// TIA Portal project "SMSS-ENLAB-01-003-1508-012-PLC-B_V13_SP1_1_V17" (V17) (continued)
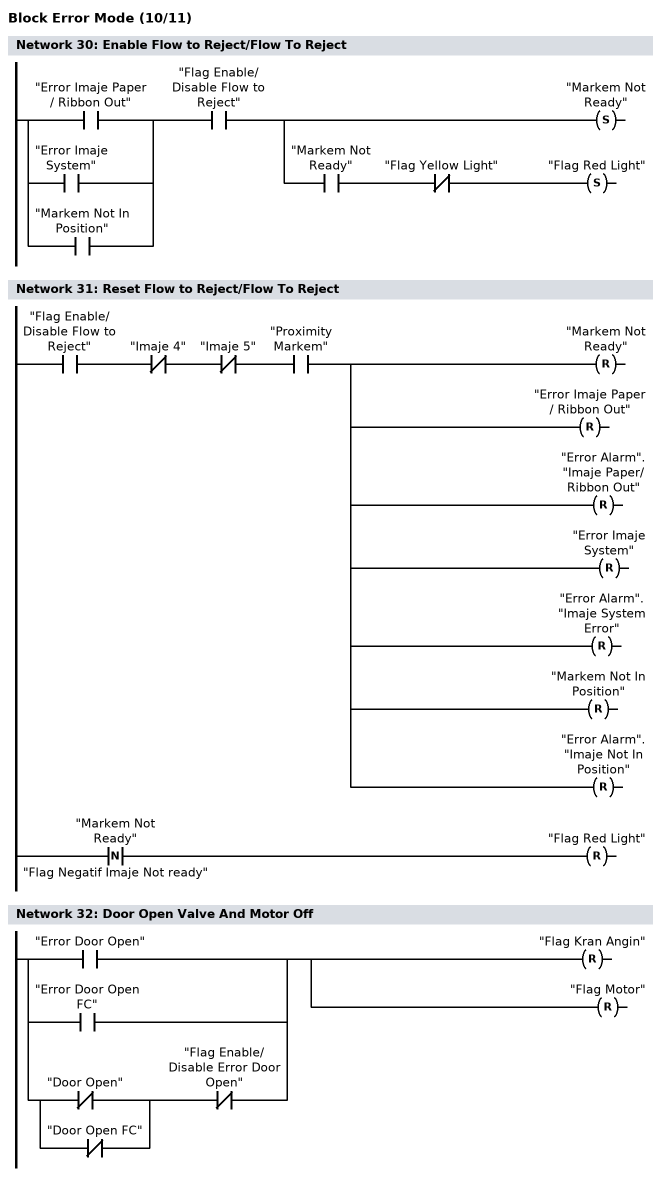
   RUNG wire#powerrail
      Contact( "Error Imaje Paper / Ribbon Out" )
      wire#w1
      Contact( "Flag Enable/Disable Flow to Reject" )
      wire#w2
      S_Coil( "Markem Not Ready" )
   END_RUNG
   RUNG wire#powerrail
      Contact( "Error Imaje System" )
   END_RUNG wire#w1
   RUNG wire#powerrail
      Contact( "Markem Not In Position" )
   END_RUNG wire#w1
   RUNG wire#w2
      Contact( "Markem Not Ready" )
      I_Contact( "Flag Yellow Light" )
      S_Coil( "Flag Red Light" )
   END_RUNG
   // the same network as SCL:
   #_w1 := ("Error Imaje Paper / Ribbon Out" OR "Error Imaje System" OR "Markem Not In Position") AND "Flag Enable/Disable Flow to Reject";
   IF #_w1 THEN "Markem Not Ready" := TRUE; END_IF;
   IF #_w1 AND "Markem Not Ready" AND NOT "Flag Yellow Light" THEN "Flag Red Light" := TRUE; END_IF;
END_REGION

REGION Network 31: Reset Flow to Reject/Flow To Reject
   RUNG wire#powerrail
      Contact( "Flag Enable/Disable Flow to Reject" )
      I_Contact( "Imaje 4" )
      I_Contact( "Imaje 5" )
      Contact( "Proximity Markem" )
      wire#w1
      R_Coil( "Markem Not Ready" )
   END_RUNG
   RUNG wire#w1
      R_Coil( "Error Imaje Paper / Ribbon Out" )
   END_RUNG
   RUNG wire#w1
      R_Coil( "Error Alarm"."Imaje Paper/Ribbon Out" )
   END_RUNG
   RUNG wire#w1
      R_Coil( "Error Imaje System" )
   END_RUNG
   RUNG wire#w1
      R_Coil( "Error Alarm"."Imaje System Error" )
   END_RUNG
   RUNG wire#w1
      R_Coil( "Markem Not In Position" )
   END_RUNG
   RUNG wire#w1
      R_Coil( "Error Alarm"."Imaje Not In Position" )
   END_RUNG
   RUNG wire#powerrail
      N_Contact(operand := "Markem Not Ready", bit := "Flag Negatif Imaje Not ready")
      R_Coil( "Flag Red Light" )
   END_RUNG
   // the same network as SCL:
   IF "Flag Enable/Disable Flow to Reject" AND NOT "Imaje 4" AND NOT "Imaje 5" AND "Proximity Markem" THEN
       "Markem Not Ready" := FALSE;
       "Error Imaje Paper / Ribbon Out" := FALSE;
       "Error Alarm"."Imaje Paper/Ribbon Out" := FALSE;
       "Error Imaje System" := FALSE;
       "Error Alarm"."Imaje System Error" := FALSE;
       "Markem Not In Position" := FALSE;
       "Error Alarm"."Imaje Not In Position" := FALSE;
   END_IF;
   #_w1 := NOT "Markem Not Ready" AND "Flag Negatif Imaje Not ready";   // falling edge of "Markem Not Ready"
   "Flag Negatif Imaje Not ready" := "Markem Not Ready";
   IF #_w1 THEN "Flag Red Light" := FALSE; END_IF;
END_REGION

REGION Network 32: Door Open Valve And Motor Off
   RUNG wire#powerrail
      Contact( "Error Door Open" )
      wire#w1
      R_Coil( "Flag Kran Angin" )
   END_RUNG
   RUNG wire#powerrail
      Contact( "Error Door Open FC" )
   END_RUNG wire#w1
   RUNG wire#powerrail
      I_Contact( "Door Open" )
      wire#w2
      I_Contact( "Flag Enable/Disable Error Door Open" )
   END_RUNG wire#w1
   RUNG wire#powerrail
      I_Contact( "Door Open FC" )
   END_RUNG wire#w2
   RUNG wire#w1
      R_Coil( "Flag Motor" )
   END_RUNG
   // the same network as SCL:
   IF "Error Door Open" OR "Error Door Open FC" OR ((NOT "Door Open" OR NOT "Door Open FC") AND NOT "Flag Enable/Disable Error Door Open") THEN
       "Flag Kran Angin" := FALSE;
       "Flag Motor" := FALSE;
   END_IF;
END_REGION

REGION Network 33: Baypas Error Reset error 3
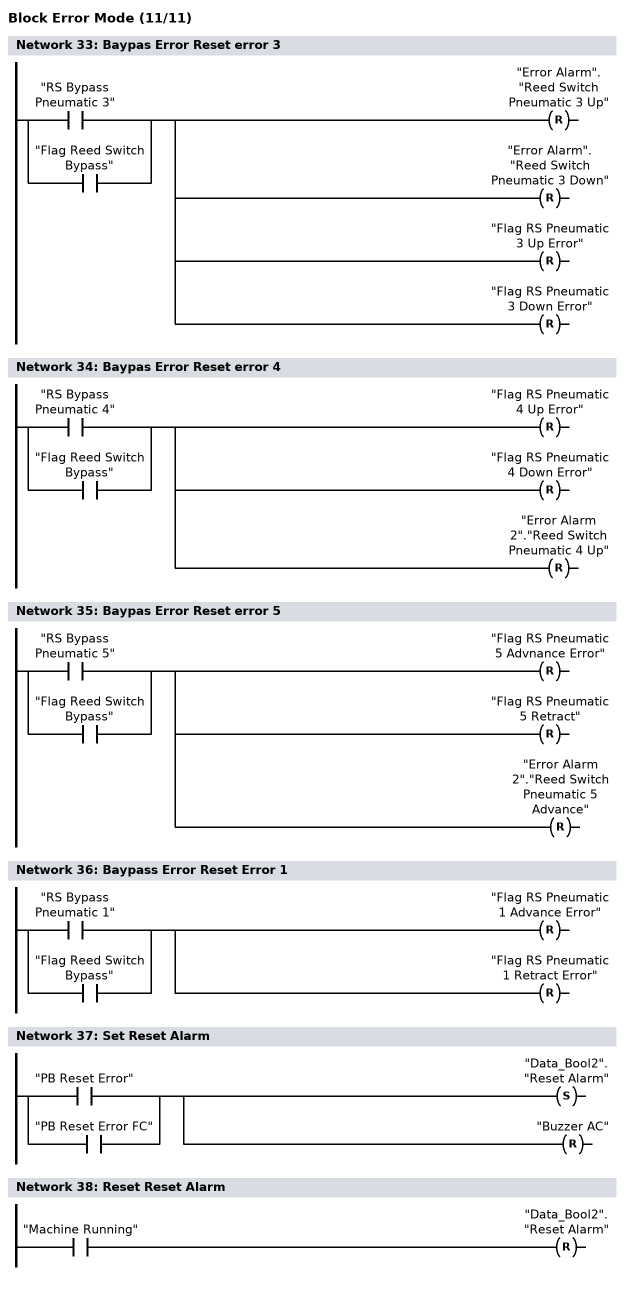
   RUNG wire#powerrail
      Contact( "RS Bypass Pneumatic 3" )
      wire#w1
      R_Coil( "Error Alarm"."Reed Switch Pneumatic 3 Up" )
   END_RUNG
   RUNG wire#powerrail
      Contact( "Flag Reed Switch Bypass" )
   END_RUNG wire#w1
   RUNG wire#w1
      R_Coil( "Error Alarm"."Reed Switch Pneumatic 3 Down" )
   END_RUNG
   RUNG wire#w1
      R_Coil( "Flag RS Pneumatic 3 Up Error" )
   END_RUNG
   RUNG wire#w1
      R_Coil( "Flag RS Pneumatic 3 Down Error" )
   END_RUNG
   // the same network as SCL:
   IF "RS Bypass Pneumatic 3" OR "Flag Reed Switch Bypass" THEN
       "Error Alarm"."Reed Switch Pneumatic 3 Up" := FALSE;
       "Error Alarm"."Reed Switch Pneumatic 3 Down" := FALSE;
       "Flag RS Pneumatic 3 Up Error" := FALSE;
       "Flag RS Pneumatic 3 Down Error" := FALSE;
   END_IF;
END_REGION

REGION Network 34: Baypas Error Reset error 4
   RUNG wire#powerrail
      Contact( "RS Bypass Pneumatic 4" )
      wire#w1
      R_Coil( "Flag RS Pneumatic 4 Up Error" )
   END_RUNG
   RUNG wire#powerrail
      Contact( "Flag Reed Switch Bypass" )
   END_RUNG wire#w1
   RUNG wire#w1
      R_Coil( "Flag RS Pneumatic 4 Down Error" )
   END_RUNG
   RUNG wire#w1
      R_Coil( "Error Alarm 2"."Reed Switch Pneumatic 4 Up" )
   END_RUNG
   // the same network as SCL:
   IF "RS Bypass Pneumatic 4" OR "Flag Reed Switch Bypass" THEN
       "Flag RS Pneumatic 4 Up Error" := FALSE;
       "Flag RS Pneumatic 4 Down Error" := FALSE;
       "Error Alarm 2"."Reed Switch Pneumatic 4 Up" := FALSE;
   END_IF;
END_REGION

REGION Network 35: Baypas Error Reset error 5
   RUNG wire#powerrail
      Contact( "RS Bypass Pneumatic 5" )
      wire#w1
      R_Coil( "Flag RS Pneumatic 5 Advnance Error" )
   END_RUNG
   RUNG wire#powerrail
      Contact( "Flag Reed Switch Bypass" )
   END_RUNG wire#w1
   RUNG wire#w1
      R_Coil( "Flag RS Pneumatic 5 Retract" )
   END_RUNG
   RUNG wire#w1
      R_Coil( "Error Alarm 2"."Reed Switch Pneumatic 5 Advance" )
   END_RUNG
   // the same network as SCL:
   IF "RS Bypass Pneumatic 5" OR "Flag Reed Switch Bypass" THEN
       "Flag RS Pneumatic 5 Advnance Error" := FALSE;
       "Flag RS Pneumatic 5 Retract" := FALSE;
       "Error Alarm 2"."Reed Switch Pneumatic 5 Advance" := FALSE;
   END_IF;
END_REGION

REGION Network 36: Baypass Error Reset Error 1
   RUNG wire#powerrail
      Contact( "RS Bypass Pneumatic 1" )
      wire#w1
      R_Coil( "Flag RS Pneumatic 1 Advance Error" )
   END_RUNG
   RUNG wire#powerrail
      Contact( "Flag Reed Switch Bypass" )
   END_RUNG wire#w1
   RUNG wire#w1
      R_Coil( "Flag RS Pneumatic 1 Retract Error" )
   END_RUNG
   // the same network as SCL:
   IF "RS Bypass Pneumatic 1" OR "Flag Reed Switch Bypass" THEN
       "Flag RS Pneumatic 1 Advance Error" := FALSE;
       "Flag RS Pneumatic 1 Retract Error" := FALSE;
   END_IF;
END_REGION

REGION Network 37: Set Reset Alarm
   RUNG wire#powerrail
      Contact( "PB Reset Error" )
      wire#w1
      S_Coil( "Data_Bool2"."Reset Alarm" )
   END_RUNG
   RUNG wire#powerrail
      Contact( "PB Reset Error FC" )
   END_RUNG wire#w1
   RUNG wire#w1
      R_Coil( "Buzzer AC" )
   END_RUNG
   // the same network as SCL:
   IF "PB Reset Error" OR "PB Reset Error FC" THEN
       "Data_Bool2"."Reset Alarm" := TRUE;
       "Buzzer AC" := FALSE;
   END_IF;
END_REGION

REGION Network 38: Reset Reset Alarm
   RUNG wire#powerrail
      Contact( "Machine Running" )
      R_Coil( "Data_Bool2"."Reset Alarm" )
   END_RUNG
   // the same network as SCL:
   IF "Machine Running" THEN "Data_Bool2"."Reset Alarm" := FALSE; END_IF;
END_REGION
END_FUNCTION_BLOCK

FUNCTION_BLOCK "Block Test Mode"   // FB2, LAD
{ S7_Optimized_Access := 'TRUE' }
VERSION : 0.1
BEGIN

REGION Network 1: Set Motor Conveyor
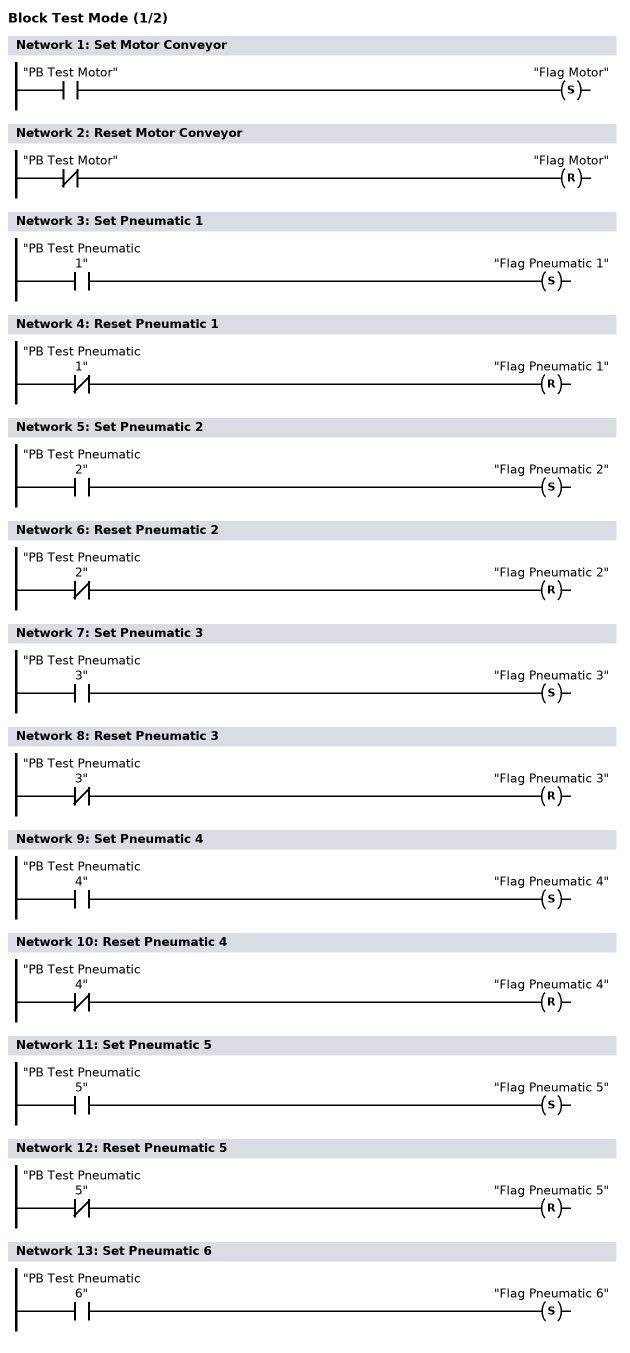
   RUNG wire#powerrail
      Contact( "PB Test Motor" )
      S_Coil( "Flag Motor" )
   END_RUNG
   // the same network as SCL:
   IF "PB Test Motor" THEN "Flag Motor" := TRUE; END_IF;
END_REGION

REGION Network 2: Reset Motor Conveyor
   RUNG wire#powerrail
      I_Contact( "PB Test Motor" )
      R_Coil( "Flag Motor" )
   END_RUNG
   // the same network as SCL:
   IF NOT "PB Test Motor" THEN "Flag Motor" := FALSE; END_IF;
END_REGION

REGION Network 3: Set Pneumatic 1
   RUNG wire#powerrail
      Contact( "PB Test Pneumatic 1" )
      S_Coil( "Flag Pneumatic 1" )
   END_RUNG
   // the same network as SCL:
   IF "PB Test Pneumatic 1" THEN "Flag Pneumatic 1" := TRUE; END_IF;
END_REGION

REGION Network 4: Reset Pneumatic 1
   RUNG wire#powerrail
      I_Contact( "PB Test Pneumatic 1" )
      R_Coil( "Flag Pneumatic 1" )
   END_RUNG
   // the same network as SCL:
   IF NOT "PB Test Pneumatic 1" THEN "Flag Pneumatic 1" := FALSE; END_IF;
END_REGION

REGION Network 5: Set Pneumatic 2
   RUNG wire#powerrail
      Contact( "PB Test Pneumatic 2" )
      S_Coil( "Flag Pneumatic 2" )
   END_RUNG
   // the same network as SCL:
   IF "PB Test Pneumatic 2" THEN "Flag Pneumatic 2" := TRUE; END_IF;
END_REGION

REGION Network 6: Reset Pneumatic 2
   RUNG wire#powerrail
      I_Contact( "PB Test Pneumatic 2" )
      R_Coil( "Flag Pneumatic 2" )
   END_RUNG
   // the same network as SCL:
   IF NOT "PB Test Pneumatic 2" THEN "Flag Pneumatic 2" := FALSE; END_IF;
END_REGION

REGION Network 7: Set Pneumatic 3
   RUNG wire#powerrail
      Contact( "PB Test Pneumatic 3" )
      S_Coil( "Flag Pneumatic 3" )
   END_RUNG
   // the same network as SCL:
   IF "PB Test Pneumatic 3" THEN "Flag Pneumatic 3" := TRUE; END_IF;
END_REGION

REGION Network 8: Reset Pneumatic 3
   RUNG wire#powerrail
      I_Contact( "PB Test Pneumatic 3" )
      R_Coil( "Flag Pneumatic 3" )
   END_RUNG
   // the same network as SCL:
   IF NOT "PB Test Pneumatic 3" THEN "Flag Pneumatic 3" := FALSE; END_IF;
END_REGION

REGION Network 9: Set Pneumatic 4
   RUNG wire#powerrail
      Contact( "PB Test Pneumatic 4" )
      S_Coil( "Flag Pneumatic 4" )
   END_RUNG
   // the same network as SCL:
   IF "PB Test Pneumatic 4" THEN "Flag Pneumatic 4" := TRUE; END_IF;
END_REGION

REGION Network 10: Reset Pneumatic 4
   RUNG wire#powerrail
      I_Contact( "PB Test Pneumatic 4" )
      R_Coil( "Flag Pneumatic 4" )
   END_RUNG
   // the same network as SCL:
   IF NOT "PB Test Pneumatic 4" THEN "Flag Pneumatic 4" := FALSE; END_IF;
END_REGION

REGION Network 11: Set Pneumatic 5
   RUNG wire#powerrail
      Contact( "PB Test Pneumatic 5" )
      S_Coil( "Flag Pneumatic 5" )
   END_RUNG
   // the same network as SCL:
   IF "PB Test Pneumatic 5" THEN "Flag Pneumatic 5" := TRUE; END_IF;
END_REGION

REGION Network 12: Reset Pneumatic 5
   RUNG wire#powerrail
      I_Contact( "PB Test Pneumatic 5" )
      R_Coil( "Flag Pneumatic 5" )
   END_RUNG
   // the same network as SCL:
   IF NOT "PB Test Pneumatic 5" THEN "Flag Pneumatic 5" := FALSE; END_IF;
END_REGION

REGION Network 13: Set Pneumatic 6
   RUNG wire#powerrail
      Contact( "PB Test Pneumatic 6" )
      S_Coil( "Flag Pneumatic 6" )
   END_RUNG
   // the same network as SCL:
   IF "PB Test Pneumatic 6" THEN "Flag Pneumatic 6" := TRUE; END_IF;
END_REGION

REGION Network 14: Reset Pneumatic 6
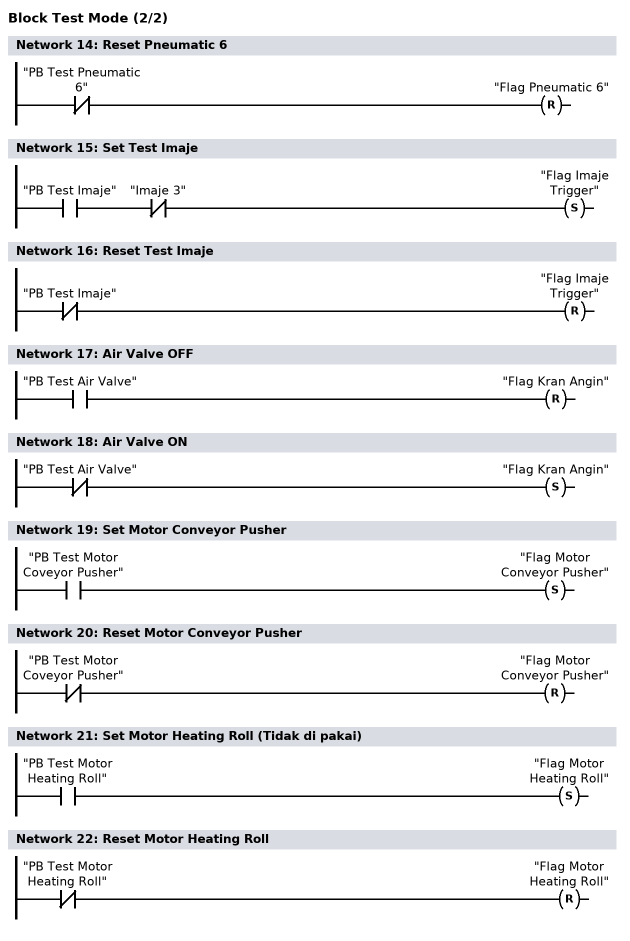
   RUNG wire#powerrail
      I_Contact( "PB Test Pneumatic 6" )
      R_Coil( "Flag Pneumatic 6" )
   END_RUNG
   // the same network as SCL:
   IF NOT "PB Test Pneumatic 6" THEN "Flag Pneumatic 6" := FALSE; END_IF;
END_REGION

REGION Network 15: Set Test Imaje
   RUNG wire#powerrail
      Contact( "PB Test Imaje" )
      I_Contact( "Imaje 3" )
      S_Coil( "Flag Imaje Trigger" )
   END_RUNG
   // the same network as SCL:
   IF "PB Test Imaje" AND NOT "Imaje 3" THEN "Flag Imaje Trigger" := TRUE; END_IF;
END_REGION

REGION Network 16: Reset Test Imaje
   RUNG wire#powerrail
      I_Contact( "PB Test Imaje" )
      R_Coil( "Flag Imaje Trigger" )
   END_RUNG
   // the same network as SCL:
   IF NOT "PB Test Imaje" THEN "Flag Imaje Trigger" := FALSE; END_IF;
END_REGION

REGION Network 17: Air Valve OFF
   RUNG wire#powerrail
      Contact( "PB Test Air Valve" )
      R_Coil( "Flag Kran Angin" )
   END_RUNG
   // the same network as SCL:
   IF "PB Test Air Valve" THEN "Flag Kran Angin" := FALSE; END_IF;
END_REGION

REGION Network 18: Air Valve ON
   RUNG wire#powerrail
      I_Contact( "PB Test Air Valve" )
      S_Coil( "Flag Kran Angin" )
   END_RUNG
   // the same network as SCL:
   IF NOT "PB Test Air Valve" THEN "Flag Kran Angin" := TRUE; END_IF;
END_REGION

REGION Network 19: Set Motor Conveyor Pusher
   RUNG wire#powerrail
      Contact( "PB Test Motor Coveyor Pusher" )
      S_Coil( "Flag Motor Conveyor Pusher" )
   END_RUNG
   // the same network as SCL:
   IF "PB Test Motor Coveyor Pusher" THEN "Flag Motor Conveyor Pusher" := TRUE; END_IF;
END_REGION

REGION Network 20: Reset Motor Conveyor Pusher
   RUNG wire#powerrail
      I_Contact( "PB Test Motor Coveyor Pusher" )
      R_Coil( "Flag Motor Conveyor Pusher" )
   END_RUNG
   // the same network as SCL:
   IF NOT "PB Test Motor Coveyor Pusher" THEN "Flag Motor Conveyor Pusher" := FALSE; END_IF;
END_REGION

REGION Network 21: Set Motor Heating Roll (Tidak di pakai)
   RUNG wire#powerrail
      Contact( "PB Test Motor Heating Roll" )
      S_Coil( "Flag Motor Heating Roll" )
   END_RUNG
   // the same network as SCL:
   IF "PB Test Motor Heating Roll" THEN "Flag Motor Heating Roll" := TRUE; END_IF;
END_REGION

REGION Network 22: Reset Motor Heating Roll
   RUNG wire#powerrail
      I_Contact( "PB Test Motor Heating Roll" )
      R_Coil( "Flag Motor Heating Roll" )
   END_RUNG
   // the same network as SCL:
   IF NOT "PB Test Motor Heating Roll" THEN "Flag Motor Heating Roll" := FALSE; END_IF;
END_REGION
END_FUNCTION_BLOCK

FUNCTION_BLOCK "Block Output"   // FB3, LAD
{ S7_Optimized_Access := 'TRUE' }
VERSION : 0.1
   VAR_TEMP   // added for the SCL form of the ladder/FBD networks
      _w1 : Bool;
      _w2 : Bool;
      _w3 : Bool;
   END_VAR
BEGIN

REGION Network 1: Red Light Tower
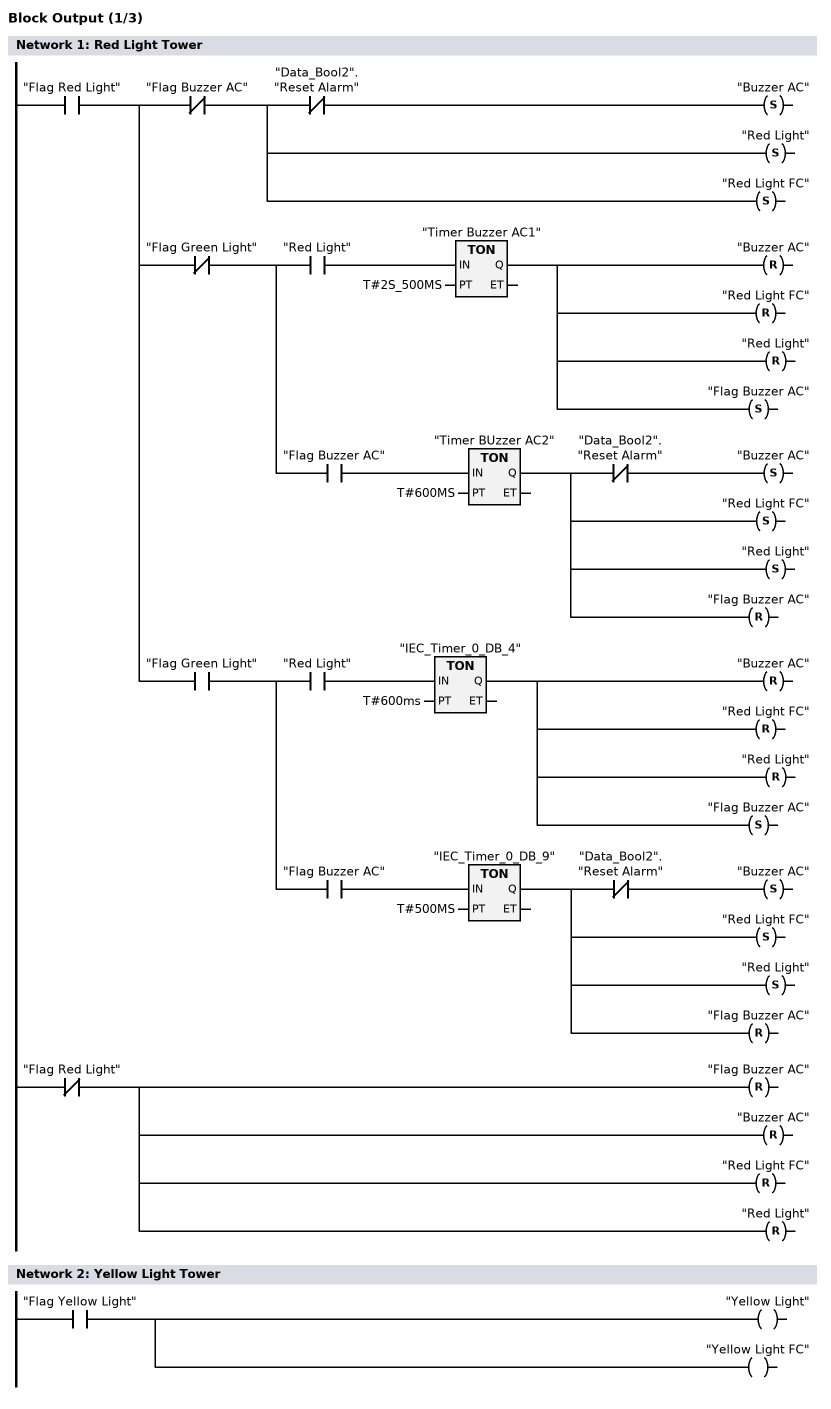
   #_w1 := "Flag Red Light" AND NOT "Flag Buzzer AC";
   IF #_w1 AND NOT "Data_Bool2"."Reset Alarm" THEN "Buzzer AC" := TRUE; END_IF;
   IF #_w1 THEN
       "Red Light" := TRUE;
       "Red Light FC" := TRUE;
   END_IF;
   #_w2 := "Flag Red Light" AND NOT "Flag Green Light";
   "Timer Buzzer AC1".TON(IN := #_w2 AND "Red Light", PT := T#2S_500MS);
   IF "Timer Buzzer AC1".Q THEN
       "Buzzer AC" := FALSE;
       "Red Light FC" := FALSE;
       "Red Light" := FALSE;
       "Flag Buzzer AC" := TRUE;
   END_IF;
   "Timer BUzzer AC2".TON(IN := #_w2 AND "Flag Buzzer AC", PT := T#600MS);
   IF "Timer BUzzer AC2".Q AND NOT "Data_Bool2"."Reset Alarm" THEN "Buzzer AC" := TRUE; END_IF;
   IF "Timer BUzzer AC2".Q THEN
       "Red Light FC" := TRUE;
       "Red Light" := TRUE;
       "Flag Buzzer AC" := FALSE;
   END_IF;
   #_w3 := "Flag Red Light" AND "Flag Green Light";
   "IEC_Timer_0_DB_4".TON(IN := #_w3 AND "Red Light", PT := T#600ms);
   IF "IEC_Timer_0_DB_4".Q THEN
       "Buzzer AC" := FALSE;
       "Red Light FC" := FALSE;
       "Red Light" := FALSE;
       "Flag Buzzer AC" := TRUE;
   END_IF;
   "IEC_Timer_0_DB_9".TON(IN := #_w3 AND "Flag Buzzer AC", PT := T#500MS);
   IF "IEC_Timer_0_DB_9".Q AND NOT "Data_Bool2"."Reset Alarm" THEN "Buzzer AC" := TRUE; END_IF;
   IF "IEC_Timer_0_DB_9".Q THEN
       "Red Light FC" := TRUE;
       "Red Light" := TRUE;
       "Flag Buzzer AC" := FALSE;
   END_IF;
   IF NOT "Flag Red Light" THEN
       "Flag Buzzer AC" := FALSE;
       "Buzzer AC" := FALSE;
       "Red Light FC" := FALSE;
       "Red Light" := FALSE;
   END_IF;
END_REGION

REGION Network 2: Yellow Light Tower
   RUNG wire#powerrail
      Contact( "Flag Yellow Light" )
      wire#w1
      Coil( "Yellow Light" )
   END_RUNG
   RUNG wire#w1
      Coil( "Yellow Light FC" )
   END_RUNG
   // the same network as SCL:
   "Yellow Light" := "Flag Yellow Light";
   "Yellow Light FC" := "Flag Yellow Light";
END_REGION

REGION Network 3: Green Light Tower
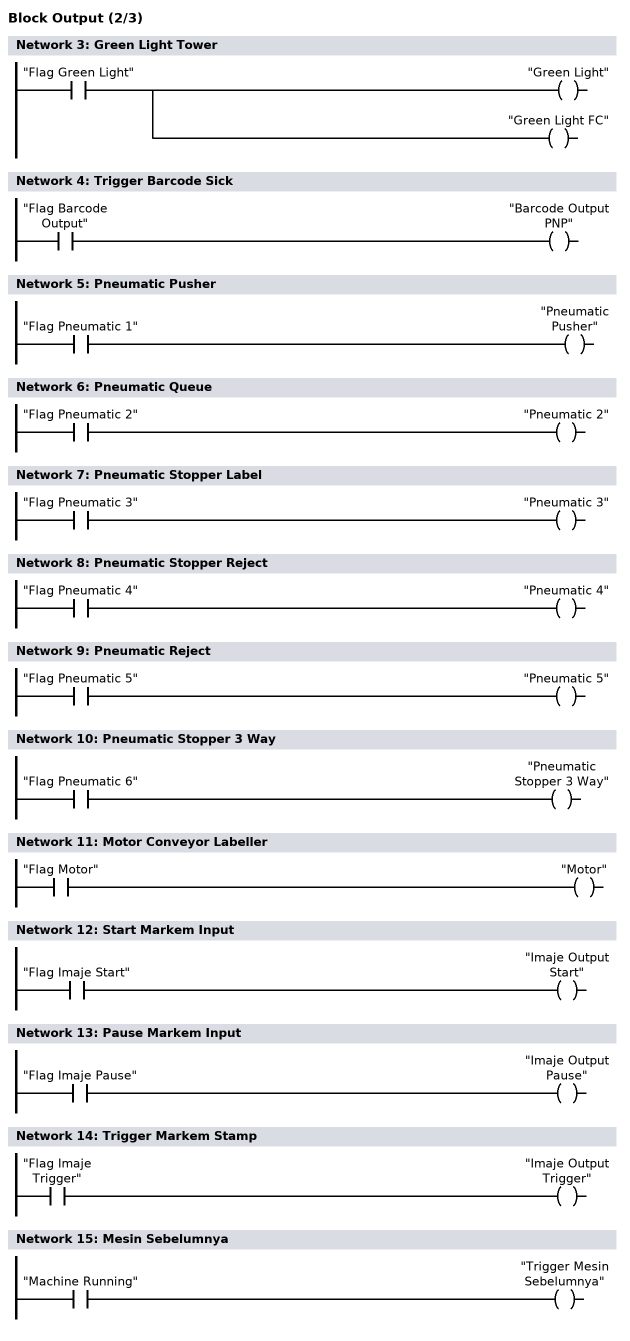
   RUNG wire#powerrail
      Contact( "Flag Green Light" )
      wire#w1
      Coil( "Green Light" )
   END_RUNG
   RUNG wire#w1
      Coil( "Green Light FC" )
   END_RUNG
   // the same network as SCL:
   "Green Light" := "Flag Green Light";
   "Green Light FC" := "Flag Green Light";
END_REGION

REGION Network 4: Trigger Barcode Sick
   RUNG wire#powerrail
      Contact( "Flag Barcode Output" )
      Coil( "Barcode Output PNP" )
   END_RUNG
   // the same network as SCL:
   "Barcode Output PNP" := "Flag Barcode Output";
END_REGION

REGION Network 5: Pneumatic Pusher
   RUNG wire#powerrail
      Contact( "Flag Pneumatic 1" )
      Coil( "Pneumatic Pusher" )
   END_RUNG
   // the same network as SCL:
   "Pneumatic Pusher" := "Flag Pneumatic 1";
END_REGION

REGION Network 6: Pneumatic Queue
   RUNG wire#powerrail
      Contact( "Flag Pneumatic 2" )
      Coil( "Pneumatic 2" )
   END_RUNG
   // the same network as SCL:
   "Pneumatic 2" := "Flag Pneumatic 2";
END_REGION

REGION Network 7: Pneumatic Stopper Label
   RUNG wire#powerrail
      Contact( "Flag Pneumatic 3" )
      Coil( "Pneumatic 3" )
   END_RUNG
   // the same network as SCL:
   "Pneumatic 3" := "Flag Pneumatic 3";
END_REGION

REGION Network 8: Pneumatic Stopper Reject
   RUNG wire#powerrail
      Contact( "Flag Pneumatic 4" )
      Coil( "Pneumatic 4" )
   END_RUNG
   // the same network as SCL:
   "Pneumatic 4" := "Flag Pneumatic 4";
END_REGION

REGION Network 9: Pneumatic Reject
   RUNG wire#powerrail
      Contact( "Flag Pneumatic 5" )
      Coil( "Pneumatic 5" )
   END_RUNG
   // the same network as SCL:
   "Pneumatic 5" := "Flag Pneumatic 5";
END_REGION

REGION Network 10: Pneumatic Stopper 3 Way
   RUNG wire#powerrail
      Contact( "Flag Pneumatic 6" )
      Coil( "Pneumatic Stopper 3 Way" )
   END_RUNG
   // the same network as SCL:
   "Pneumatic Stopper 3 Way" := "Flag Pneumatic 6";
END_REGION

